HMI tags "Default tag table"
   "66_Event_Data_BC_EVENT_WORD_01" : Word = PLC "66_Event_Data".BC_EVENT_WORD_01 AT %DB66.DBW0, 1 s
   "66_Event_Data_BC_EVENT_WORD_02" : Word = PLC "66_Event_Data".BC_EVENT_WORD_02 AT %DB66.DBW2, 1 s
   "64_Message_Data_BC_MESSAGE_WORD_01" : Word = PLC "64_Message_Data".BC_MESSAGE_WORD_01 AT %DB64.DBW0, 1 s
   "64_Message_Data_BC_MESSAGE_WORD_02" : Word = PLC "64_Message_Data".BC_MESSAGE_WORD_02 AT %DB64.DBW2, 1 s
   "66_Event_Data_IGG_EVENT_WORD_01" : Word = PLC "66_Event_Data".IGG_EVENT_WORD_01 AT %DB66.DBW0, 1 s
   "66_Event_Data_IGG_EVENT_WORD_02" : Word = PLC "66_Event_Data".IGG_EVENT_WORD_02 AT %DB66.DBW2, 1 s
   "64_Message_Data_IGG_MESSAGE_WORD_01" : Word = PLC "64_Message_Data".IGG_MESSAGE_WORD_01 AT %DB64.DBW0, 1 s
   "64_Message_Data_IGG_MESSAGE_WORD_02" : Word = PLC "64_Message_Data".IGG_MESSAGE_WORD_02 AT %DB64.DBW2, 1 s
   "Current User" : WString[15] AT %DB1.DBX0.0
   "db_time_sync_time_system_READ" : LDT = PLC db_time_sync_time_system_READ AT %M2.0, 1 s
   "80_From_HMI_Cooling System Overrun" : Time = PLC "80_From_HMI"."Cooling System Overrun", 1 s
   "Start Sequenc_DB_Post Purge Time Sec" : Int, internal
   "db_time_sync_time_local_READ" : LDT = PLC db_time_sync_time_local_READ AT %M4.0, 1 s
   "82_To_HMI_Fuel Pump 1 Animation" : Int = PLC "82_To_HMI"."Fuel Pump 1 Animation", 1 s
   "82_To_HMI_Fuel Pump 2 Animation" : Int = PLC "82_To_HMI"."Fuel Pump 2 Animation", 1 s
   "16_AQ_Data_CV203_CNTRL(1)" : Real = PLC "16_AQ_Data".CV203_CNTRL, 1 s
   "HMI Data_O2 Setpoint" : Real, internal
   "82_To_HMI_IA Compressor Animation" : Int = PLC "82_To_HMI"."IA Compressor Animation", 1 s
   "Atomising Air  Valve Manual Regulator" : Int, internal
   "Fuel Valve Manual Regulator" : Int, internal
   "82_To_HMI_I&A Compressor Run Hours(1)" : Int = PLC "82_To_HMI"."I&A Compressor Run Hours", 1 s
   "82_To_HMI_I&A Compressor Service Time Hours" : Int = PLC "82_To_HMI"."I&A Compressor Service Time Hours", 1 s
   "82_To_HMI_CA Blower Run Days" : Int = PLC "82_To_HMI"."CA Blower Run Days", 1 s
   "82_To_HMI_CA Blower Service Time Hours" : Int = PLC "82_To_HMI"."CA Blower Service Time Hours", 1 s
   "82_To_HMI_CA Blower Run Hours" : Int = PLC "82_To_HMI"."CA Blower Run Hours", 1 s
   "82_To_HMI_CA Blower Run Minutes" : Int = PLC "82_To_HMI"."CA Blower Run Minutes", 1 s
   "82_To_HMI_I&A Compressor Run Minutes" : Int = PLC "82_To_HMI"."I&A Compressor Run Minutes", 1 s
   "82_To_HMI_I&A Compressor Run Seconds" : Int = PLC "82_To_HMI"."I&A Compressor Run Seconds", 1 s
   "P305_Functioning Hours_IDB_Hours Total" : Int = PLC "P305_Functioning Hours_IDB"."Hours Total", 1 s
   "82_To_HMI_P305 FW Pump Service Time Hours" : Int = PLC "82_To_HMI"."P305 FW Pump Service Time Hours", 1 s
   "P305_Functioning Hours_IDB_Service Time bit" : Bool = PLC "P305_Functioning Hours_IDB"."Service Time bit", 1 s
   "P305_Functioning Hours_IDB_Minutes" : Int = PLC "P305_Functioning Hours_IDB".Minutes, 1 s
   "P305_Functioning Hours_IDB_Seconds" : Int = PLC "20_TANKS_IP_DATA".RIO_04.SECOND_TANK.BWT_LEVEL_HIHI, 1 s
   "FW Pump Animation" : Int, internal
   "82_To_HMI_I&A Compressor Run Hours" : Int = PLC "82_To_HMI"."I&A Compressor Run Hours", 1 s
   "82_To_HMI_CRNT_MODE_IGG" : Int = PLC "82_To_HMI".CRNT_MODE_IGG, 1 s
   "70_Mode_Data_AUT_RST_PLS_IN" : Bool = PLC "70_Mode_Data".AUT_RST_PLS.IN, 1 s
   "RESET_STEP" : Bool = PLC RESET_STEP AT %M12.0, 1 s
   "100_IGG_AUTO_SEQ_DB_CRNT_STEP" : Int = PLC "100_IGG_AUTO_SEQ_DB".CRNT_STEP, 1 s
   "100_BC_AUTO_SEQ_DB_CRNT_STEP" : Int = PLC "100_BC_AUTO_SEQ_DB".CRNT_STEP, 1 s
   "103_Main_Burner_DB_RUN" : Bool = PLC "103_Main_Burner_DB".RUN, 1 s
   "60_Alarm_Data_ALRM_PRSNT" : Bool = PLC "60_Alarm_Data".ALRM_PRSNT AT %DB60.DBX32.0, 1 s
      on ChangeValue: "ALARM_Present"()
   "62_Warning_Data_WRNG_PRSNT" : Bool = PLC "62_Warning_Data".WRNG_PRSNT AT %DB62.DBX16.0, 1 s
   "103_Main_Burner_DB_RUNNING" : Bool = PLC "103_Main_Burner_DB".RUNNING, 1 s
   "101_Fuel_Pumps_DB_Duty Is B" : Bool = PLC "101_Fuel_Pumps_DB"."Duty Is B", 1 s
   "101_Fuel_Pumps_DB_Duty Is A" : Bool = PLC "101_Fuel_Pumps_DB"."Duty Is A", 1 s
   "84_Setpoints_PIT204_High" : Real = PLC "84_Setpoints".PIT204_High, 1 s
   "84_Setpoints_PIT204_High(1)" : Real = PLC "84_Setpoints".PIT204_High, 1 s
   "84_Setpoints_PIT204_HighHigh" : Real = PLC "84_Setpoints".PIT204_HighHigh, 1 s
   "84_Setpoints_PIT204_HighHigh(1)" : Real = PLC "84_Setpoints".PIT204_HighHigh, 1 s
   "84_Setpoints_PIT204_LowLow" : Real = PLC "84_Setpoints".PIT204_LowLow, 1 s
   "84_Setpoints_PIT204_LowLow(1)" : Real = PLC "84_Setpoints".PIT204_LowLow, 1 s
   "84_Setpoints_PIT204_Low" : Real = PLC "84_Setpoints".PIT204_Low, 1 s
   "84_Setpoints_PIT204_Low(1)" : Real = PLC "84_Setpoints".PIT204_Low, 1 s
   "80_From_HMI_RST_LOCKOUT" : Bool = PLC "80_From_HMI".RST_LOCKOUT, 1 s
   "80_From_HMI_Beacon frequency" : Time = PLC "80_From_HMI"."Beacon frequency", 1 s
   "80_From_HMI_Buzzer reset time" : Time = PLC "80_From_HMI"."Buzzer reset time", 1 s
   "80_From_HMI_Reset_Alarms" : Bool = PLC "80_From_HMI".Reset_Alarms, 1 s
   "Alarm beacon handling_DB_Buzzer_Timer_0_Instance_Q" : Bool = PLC "Alarm beacon handling_DB".Buzzer_Timer_0_Instance.Q, 1 s
   "Buzzer" : Bool = PLC Buzzer AT %Q1.7, 1 s
   "80_From_HMI_FLM_FAIL_DLY" : Time = PLC "80_From_HMI".FLM_FAIL_DLY, 1 s
   "103_Main_Burner_DB_DN_OK" : Bool = PLC "103_Main_Burner_DB".DN_OK, 1 s
   "103_Main_Burner_DB_Days burn_CV" : Int = PLC "103_Main_Burner_DB"."Days burn".CV, 1 s
   "103_Main_Burner_DB_Hours burn_CV" : Int = PLC "103_Main_Burner_DB"."Hours burn".CV, 1 s
   "103_Main_Burner_DB_Minutes burn_CV" : Int = PLC "103_Main_Burner_DB"."Minutes burn".CV, 1 s
   "103_Main_Burner_DB_Seconds burn_CV" : Int = PLC "103_Main_Burner_DB"."Seconds burn".CV, 1 s
   "103_Main_Burner_DB_STATE" : Int = PLC "103_Main_Burner_DB".STATE, 1 s
   "19_AUTO_CMNDS_Data_CV203_RAMP_CNTRL" : Bool = PLC "19_AUTO_CMNDS_Data".CV203_RAMP_CNTRL, 1 s
   "102_Pilot_Burner_DB_RUNNING" : Bool = PLC "102_Pilot_Burner_DB".RUNNING, 1 s
   "68_Sys_Status_Data_FUEL_PRES_IN_RNG" : Bool = PLC "68_Sys_Status_Data".FUEL_PRES_IN_RNG, 1 s
   "68_Sys_Status_Data_IA_PRES_IN_RNG" : Bool = PLC "68_Sys_Status_Data".IA_PRES_IN_RNG, 1 s
   "84_Setpoints_Gain" : Real = PLC "84_Setpoints".Gain, 1 s
   "84_Setpoints_Integration Time" : Time = PLC "84_Setpoints"."Integration Time", 1 s
   "84_Setpoints_Derive Time" : Time = PLC "84_Setpoints"."Derive Time", 1 s
   "O2 Ramp Control_QLMN_HLM" : Bool = PLC "O2 Ramp Control".QLMN_HLM, 1 s
   "O2 Ramp Control_QLMN_LLM" : Bool = PLC "O2 Ramp Control".QLMN_LLM, 1 s
   "84_Setpoints_P_ON" : Bool = PLC "84_Setpoints".P_ON, 1 s
   "84_Setpoints_I_ON" : Bool = PLC "84_Setpoints".I_ON, 1 s
   "84_Setpoints_D_ON" : Bool = PLC "84_Setpoints".D_ON, 1 s
   "Evolving Setpoint_DB_LevelBetter" : Bool = PLC "Evolving Setpoint_DB".LevelBetter, 1 s
   "84_Setpoints_Max Opening" : Real = PLC "84_Setpoints"."Max Opening", 1 s
   "84_Setpoints_Min Opening" : Real = PLC "86_Times".STEP_MAX_TIME_STP_290, 1 s
   "80_From_HMI_Post Purge Time" : Time = PLC "80_From_HMI"."Post Purge Time", 1 s
   "103_Main_Burner_DB_Status" : Int = PLC "103_Main_Burner_DB".Status, 1 s
   "80_From_HMI_Reset CV203 PID" : Bool = PLC "80_From_HMI"."Reset CV203 PID", 1 s
   "80_From_HMI_BurnerProgramedStop" : Bool = PLC "80_From_HMI".BurnerProgramedStop, 1 s
   "82_To_HMI_CA Blower Reset Hours" : Bool = PLC "82_To_HMI"."CA Blower Reset Hours", 1 s
   "82_To_HMI_CA Blower Service Due" : Bool = PLC "82_To_HMI"."CA Blower Service Due", 1 s
   "Operation hours E139_IDB_Hours Functioning" : Int = PLC "Operation hours E139_IDB"."Hours Functioning", 1 s
   "82_To_HMI_CA Blower Total Run Hours" : Int = PLC "82_To_HMI"."CA Blower Total Run Hours", 1 s
   "82_To_HMI_I&A Compressor Total Run Hours" : Int = PLC "82_To_HMI"."I&A Compressor Total Run Hours", 1 s
   "82_To_HMI_I&A Compressor Reset Hours" : Bool = PLC "82_To_HMI"."I&A Compressor Reset Hours", 1 s
   "82_To_HMI_I&A Compressor Service Due" : Bool = PLC "82_To_HMI"."I&A Compressor Service Due", 1 s
   "82_To_HMI_E500A Fuel Pump Run Hours" : Int = PLC "82_To_HMI"."E500A Fuel Pump Run Hours", 1 s
   "64_Functioning Hours_E500A_IDB_Hours Functioning" : Int = PLC "64_Functioning Hours_E500A_IDB"."Hours Functioning", 1 s
   "82_To_HMI_E500A Fuel Pump Run Minutes" : Int = PLC "82_To_HMI"."E500A Fuel Pump Run Minutes", 1 s
   "82_To_HMI_E500A Fuel Pump Run Seconds" : Int = PLC "82_To_HMI"."E500A Fuel Pump Run Seconds", 1 s
   "82_To_HMI_E500A Fuel Pump Total Run Hours" : Int = PLC "82_To_HMI"."E500A Fuel Pump Total Run Hours", 1 s
   "82_To_HMI_E500A Fuel Pump Service Time Hours" : Int = PLC "82_To_HMI"."E500A Fuel Pump Service Time Hours", 1 s
   "82_To_HMI_E500A Fuel Pump Reset Hours" : Bool = PLC "82_To_HMI"."E500A Fuel Pump Reset Hours", 1 s
   "64_Functioning Hours_E500B_IDB_Hours Functioning" : Int = PLC "64_Functioning Hours_E500B_IDB"."Hours Functioning", 1 s
   "82_To_HMI_E500B Fuel Pump Run Minutes" : Int = PLC "82_To_HMI"."E500B Fuel Pump Run Minutes", 1 s
   "82_To_HMI_E500B Fuel Pump Run Seconds" : Int = PLC "82_To_HMI"."E500B Fuel Pump Run Seconds", 1 s
   "82_To_HMI_E500B Fuel Pump Total Run Hours" : Int = PLC "82_To_HMI"."E500B Fuel Pump Total Run Hours", 1 s
   "82_To_HMI_E500B Fuel Pump Service Time Hours" : Int = PLC "82_To_HMI"."E500B Fuel Pump Service Time Hours", 1 s
   "82_To_HMI_E500B Fuel Pump Reset Hours" : Bool = PLC "82_To_HMI"."E500B Fuel Pump Reset Hours", 1 s
   "82_To_HMI_E500B Fuel Pump Service Due" : Bool = PLC "82_To_HMI"."E500B Fuel Pump Service Due", 1 s
   "82_To_HMI_E500A Fuel Pump Service Due" : Bool = PLC "82_To_HMI"."E500A Fuel Pump Service Due", 1 s
   "64_Functioning Hours_P301_IDB_Hours Functioning" : Int = PLC "64_Functioning Hours_P301_IDB"."Hours Functioning", 1 s
   "82_To_HMI_P301 CSW Pump Run Minutes" : Int = PLC "82_To_HMI"."P301 CSW Pump Run Minutes", 1 s
   "82_To_HMI_P301 CSW Pump Run Seconds" : Int = PLC "82_To_HMI"."P301 CSW Pump Run Seconds", 1 s
   "82_To_HMI_P301 CSW Pump Reset Hours" : Bool = PLC "82_To_HMI"."P301 CSW Pump Reset Hours", 1 s
   "82_To_HMI_P301 CSW Pump Service Due" : Bool = PLC "82_To_HMI"."P301 CSW Pump Service Due", 1 s
   "80_From_HMI_P301_PRSNT" : Bool = PLC "80_From_HMI".P301_PRSNT, 1 s
   "Alarms_Acknowledge_IGG_ALARM_ACKNLG_3" : Word = PLC Alarms_Acknowledge.IGG_ALARM_ACKNLG_3 AT %DB67.DBW4, 1 s
   "Alarms_Acknowledge_IGG_ALARM_ACKNLG_4" : Word = PLC Alarms_Acknowledge.IGG_ALARM_ACKNLG_4 AT %DB67.DBW6, 1 s
   "Alarms_Acknowledge_IGG_ALARM_ACKNLG_2" : Word = PLC Alarms_Acknowledge.IGG_ALARM_ACKNLG_2 AT %DB67.DBW2, 1 s
   "Alarms_Acknowledge_IGG_ALARM_ACKNLG_1" : Word = PLC Alarms_Acknowledge.IGG_ALARM_ACKNLG_1 AT %DB67.DBW0, 1 s
   "BC_ALARM_ACKNLG_1" : Word = PLC BC_ALARM_ACKNLG_1 AT %MW24, 1 s
   "BC_ALARM_ACKNLG_2" : Word = PLC BC_ALARM_ACKNLG_2 AT %MW26, 1 s
   "BC_ALARM_ACKNLG_3" : Word = PLC BC_ALARM_ACKNLG_3 AT %MW28, 1 s
   "BC_ALARM_ACKNLG_4" : Word = PLC BC_ALARM_ACKNLG_4 AT %MW30, 1 s
   "80_From_HMI_P305_PRSNT" : Bool = PLC "80_From_HMI".P305_PRSNT, 1 s
   "68_Sys_Status_Data_INTRLKS_OK" : Bool = PLC "68_Sys_Status_Data".INTRLKS_OK, 1 s
   "82_To_HMI_E-STOP LATCHED" : Bool = PLC "82_To_HMI"."E-STOP LATCHED", 1 s
   "82_To_HMI_P301 CSW Pump Run Days" : Int = PLC "82_To_HMI"."P301 CSW Pump Run Days", 1 s
   "82_To_HMI_CA Blower Run Seconds" : Int = PLC "82_To_HMI"."CA Blower Run Seconds", 1 s
   "82_To_HMI_P305 FW Pump Reset Hours" : Bool = PLC "82_To_HMI"."P305 FW Pump Reset Hours", 1 s
   "P305_Functioning Hours_IDB_Hours Functioning Out" : Int = PLC "P305_Functioning Hours_IDB"."Hours Functioning Out", 1 s
   "82_To_HMI_P305 FW Pump Run Hours" : Int = PLC "82_To_HMI"."P305 FW Pump Run Hours", 1 s
   "82_To_HMI_P305 FW Pump Run Days" : Int = PLC "82_To_HMI"."P305 FW Pump Run Days", 1 s
   "82_To_HMI_P301 CSW Pump Service Time Hours" : Int = PLC "82_To_HMI"."P301 CSW Pump Service Time Hours", 1 s
   "82_To_HMI_P301 CSW Pump Run Hours" : Int = PLC "82_To_HMI"."P301 CSW Pump Run Hours", 1 s
   "82_To_HMI_P301 CSW Pump Total Run Hours" : Int = PLC "82_To_HMI"."P301 CSW Pump Total Run Hours", 1 s
   "80_From_HMI_PIT 359 delay" : Time = PLC "80_From_HMI"."PIT 359 delay", 1 s
   "80_From_HMI_PIT 316 delay" : Time = PLC "80_From_HMI"."PIT 316 delay", 1 s
   "86_Times_PIT353 Delay" : Time = PLC "86_Times"."PIT353 Delay", 1 s
   "86_Times_PIT416 Delay" : Time = PLC "86_Times"."PIT416 Delay", 1 s
   "19_AUTO_CMNDS_Data_PIT416_CMND_Target" : Real = PLC "19_AUTO_CMNDS_Data".PIT416_CMND_Target, 1 s
   "2102_TIME_CALCS_DB_Voyage_TIME_days" : Int = PLC "2102_TIME_CALCS_DB".Voyage_TIME_days, 1 s
   "2102_TIME_CALCS_DB_Voyage_TIME_invalid" : Bool = PLC "2102_TIME_CALCS_DB".Voyage_TIME_invalid AT %DB1.DBW0, 1 s
      on ChangeValue: "VoyageTimeInsufficient"()
   "2102_TIME_CALCS_DB_TOT_SEQ_DAYS" : Real = PLC "2102_TIME_CALCS_DB".TOT_SEQ_DAYS, 1 s
   "2102_TIME_CALCS_DB_POST_DWELL_TMR_DN(1)" : Bool = PLC "2102_TIME_CALCS_DB".POST_DWELL_TMR_DN AT %DB1.DBD0, 1 s
   "2102_TIME_CALCS_DB_PRE-DWEL HOURS REMNG" : Int = PLC "2102_TIME_CALCS_DB"."PRE-DWEL HOURS REMNG" AT %DB1.DBW0, 1 s
   "504_Tank Grouping_DB2020_TANK ACTIV 2" : Bool = PLC "504_Tank Grouping_DB2020"."TANK ACTIV 2" AT %DB1.DBW0, 1 s
   "504_Tank Grouping_DB2020_TANK ACTIV 4" : Bool = PLC "504_Tank Grouping_DB2020"."TANK ACTIV 4" AT %DB1.DBW0, 1 s
   "504_Tank Grouping_DB2020_TANK ACTIV 6" : Bool = PLC "504_Tank Grouping_DB2020"."TANK ACTIV 6" AT %DB1.DBW0, 1 s
   "504_Tank Grouping_DB2020_TANK ACTIV 8" : Bool = PLC "504_Tank Grouping_DB2020"."TANK ACTIV 8" AT %DB1.DBW0, 1 s
   "504_Tank Grouping_DB2020_TANK ACTIV 10" : Bool = PLC "504_Tank Grouping_DB2020"."TANK ACTIV 10" AT %DB1.DBW0, 1 s
   "504_Tank Grouping_DB2020_TANK ACTIV 12" : Bool = PLC "504_Tank Grouping_DB2020"."TANK ACTIV 12" AT %DB1.DBW0, 1 s
   "504_Tank Grouping_DB2020_TANK ACTIV 14" : Bool = PLC "504_Tank Grouping_DB2020"."TANK ACTIV 14" AT %DB1.DBW0, 1 s
   "504_Tank Grouping_DB2020_TANK ACTIV 16" : Bool = PLC "504_Tank Grouping_DB2020"."TANK ACTIV 16" AT %DB1.DBW0, 1 s
   "504_Tank Grouping_DB2020_TANK ACTIV 18" : Bool = PLC "504_Tank Grouping_DB2020"."TANK ACTIV 18" AT %DB1.DBW0, 1 s
   "504_Tank Grouping_DB2020_TANK ACTIV 20" : Bool = PLC "504_Tank Grouping_DB2020"."TANK ACTIV 20" AT %DB1.DBW0, 1 s
   "504_Tank Grouping_DB2020_TANK ACTIV 3" : Bool = PLC "504_Tank Grouping_DB2020"."TANK ACTIV 3" AT %DB1.DBW0, 1 s
   "504_Tank Grouping_DB2020_TANK ACTIV 5" : Bool = PLC "504_Tank Grouping_DB2020"."TANK ACTIV 5" AT %DB1.DBW0, 1 s
   "504_Tank Grouping_DB2020_TANK ACTIV 7" : Bool = PLC "504_Tank Grouping_DB2020"."TANK ACTIV 7" AT %DB1.DBW0, 1 s
   "504_Tank Grouping_DB2020_TANK ACTIV 9" : Bool = PLC "504_Tank Grouping_DB2020"."TANK ACTIV 9" AT %DB1.DBW0, 1 s
   "504_Tank Grouping_DB2020_TANK ACTIV 11" : Bool = PLC "504_Tank Grouping_DB2020"."TANK ACTIV 11" AT %DB1.DBW0, 1 s
   "504_Tank Grouping_DB2020_TANK ACTIV 13" : Bool = PLC "504_Tank Grouping_DB2020"."TANK ACTIV 13" AT %DB1.DBW0, 1 s
   "504_Tank Grouping_DB2020_TANK ACTIV 1" : Bool = PLC "504_Tank Grouping_DB2020"."TANK ACTIV 1" AT %DB1.DBW0, 1 s
   "504_Tank Grouping_DB2020_TANK ACTIV 17" : Bool = PLC "504_Tank Grouping_DB2020"."TANK ACTIV 17" AT %DB1.DBW0, 1 s
   "504_Tank Grouping_DB2020_TANK ACTIV 19" : Bool = PLC "504_Tank Grouping_DB2020"."TANK ACTIV 19" AT %DB1.DBW0, 1 s
   "504_Tank Grouping_DB2020_TANK ACTIV 21" : Bool = PLC "504_Tank Grouping_DB2020"."TANK ACTIV 21" AT %DB1.DBW0, 1 s
   "2110_BTCS_CNTRL_DB_PORT_TANK_STS(1)" : Bool = PLC "2110_BTCS_CNTRL_DB".PORT_TANK_STS AT %DB1.DBX0.0, 1 s
   "Tank Activated Port 2" : Int, internal
   "Tank Activated Port 3" : Int, internal
   "Tank Activated Port 4" : Int, internal
   "Tank Activated Port 5" : Int, internal
   "Tank Activated Port 6" : Int, internal
   "Tank Activated Port 7" : Int, internal
   "Tank Activated Port 8" : Int, internal
   "Tank Activated Port 9" : Int, internal
   "Tank Activated Port 10" : Int, internal
   "2110_BTCS_CNTRL_DB_STBD_TANK_STS(1)" : Bool = PLC "20_TANKS_IP_DATA".RIO_01.FIRST_TANK.GTT_ISOL_VALVE_OPEN, 1 s
   "Tank Activated Star 2" : Int, internal
   "Tank Activated Star 3" : Int, internal
   "Tank Activated Star 4" : Int, internal
   "Tank Activated Star 5" : Int, internal
   "Tank Activated Star 6" : Int, internal
   "Tank Activated Star 7" : Int, internal
   "Tank Activated Star 8" : Int, internal
   "Tank Activated Star 9" : Int, internal
   "Tank Activated Star 10" : Int, internal
   "2102_TIME_CALCS_DB_PRE-DWEL_Warning 1" : Bool = PLC "2102_TIME_CALCS_DB"."PRE-DWEL_Warning 1", 500 ms
      on ChangeValue: "TimeRemainingToTreatment"()
   "2102_TIME_CALCS_DB_PRE-DWEL_Warning Min 1" : Int = PLC "2102_TIME_CALCS_DB"."PRE-DWEL_Warning Min 1", 1 s
   "2102_TIME_CALCS_DB_PRE-DWEL_Warning Min 2" : Int = PLC "2102_TIME_CALCS_DB"."PRE-DWEL_Warning Min 2", 1 s
   "2102_TIME_CALCS_DB_PRE-DWEL_Warning Min 3" : Int = PLC "2102_TIME_CALCS_DB"."PRE-DWEL_Warning Min 3", 1 s
   "2102_TIME_CALCS_DB_PRE-DWEL_Warning Reset 1" : Bool = PLC "2102_TIME_CALCS_DB"."PRE-DWEL_Warning Reset 1", 1 s
   "2102_TIME_CALCS_DB_PRE-DWEL_Warning 2" : Bool = PLC "2102_TIME_CALCS_DB"."PRE-DWEL_Warning 2", 500 ms
      on ChangeValue: "TreatmentRequired"()
   "2102_TIME_CALCS_DB_PRE-DWEL_Warning 3" : Bool = PLC "2102_TIME_CALCS_DB"."PRE-DWEL_Warning 3", 1 s
   "2102_TIME_CALCS_DB_PRE-DWEL_Warning Reset 2" : Bool = PLC "2102_TIME_CALCS_DB"."PRE-DWEL_Warning Reset 2", 1 s
   "2102_TIME_CALCS_DB_PRE-DWEL_Warning Reset 3" : Bool = PLC "2102_TIME_CALCS_DB"."PRE-DWEL_Warning Reset 3", 1 s
   "2102_TIME_CALCS_DB_60X boost" : Bool = PLC "2102_TIME_CALCS_DB"."60X boost", 1 s
   "86_Times_P301_START_DLY" : Time = PLC "86_Times".P301_START_DLY, 1 s
   "86_Times_FS332 Delay" : Time = PLC "86_Times"."FS332 Delay", 1 s
   "86_Times_LIT304 Delay" : Time = PLC "86_Times"."LIT304 Delay", 1 s
   "86_Times_PIT402_Ramp_Seconds" : Int = PLC "86_Times".PIT402_Ramp_Seconds, 1 s
   "86_Times_PIT402 Alarm Delay" : Time = PLC "86_Times"."PIT402 Alarm Delay", 1 s
   "84_Setpoints_PIT113_Burner_Target" : Real = PLC "84_Setpoints".PIT113_Burner_Target, 1 s
   "2102_TIME_CALCS_DB_PRE-DWEL MINS REMNG" : Int = PLC "2102_TIME_CALCS_DB"."PRE-DWEL MINS REMNG", 1 s
   "84_Setpoints_LIT304_InitialFill_Target_Low" : Real = PLC "84_Setpoints".LIT304_InitialFill_Target_Low, 1 s
   "84_Setpoints_LIT304_Refill_Target_Low" : Real = PLC "84_Setpoints".LIT304_Refill_Target_Low, 1 s
   "1111_PID_CV111_Setpoint" : Real = PLC "1111_PID_CV111".Setpoint, 1 s
   "2086_Times_TT426_PORT_Alarm Delay" : Time = PLC "2086_Times"."TT426_PORT_Alarm Delay", 1 s
   "2086_Times_TT426_STAR_Alarm Delay" : Time = PLC "2086_Times"."TT426_STAR_Alarm Delay", 1 s
   "2086_Times_FIT418PORT Alarm Delay" : Time = PLC "2086_Times"."FIT418PORT Alarm Delay", 1 s
   "2086_Times_FIT420PORT Alarm Delay" : Time = PLC "2086_Times"."FIT420PORT Alarm Delay", 1 s
   "2086_Times_FIT417STAR Alarm Delay" : Time = PLC "2086_Times"."FIT417STAR Alarm Delay", 1 s
   "2086_Times_FIT419STAR Alarm Delay" : Time = PLC "2086_Times"."FIT419STAR Alarm Delay", 1 s
   "2086_Times_PT415 Alarm Delay" : Time = PLC "2086_Times"."PT415 Alarm Delay", 1 s
   "2086_Times_PIT424 Alarm Delay" : Time = PLC "2086_Times"."PIT424 Alarm Delay", 1 s
   "2086_Times_LS425 Port Alarm Delay" : Time = PLC "2086_Times"."LS425 Port Alarm Delay", 1 s
   "2086_Times_LS425 Star Alarm Delay" : Time = PLC "2086_Times"."LS425 Star Alarm Delay", 1 s
   "2086_Times_PS436 Alarm Delay" : Time = PLC "2086_Times"."PS436 Alarm Delay", 1 s
   "2102_TIME_CALCS_DB_Voyage_TIME_remaining_m" : Int = PLC "2102_TIME_CALCS_DB".Voyage_TIME_remaining_m, 1 s
   "2102_TIME_CALCS_DB_Voyage_TIME_remaining_h" : Int = PLC "2102_TIME_CALCS_DB".Voyage_TIME_remaining_h, 1 s
   "2102_TIME_CALCS_DB_Time_To_Treatment" : Int = PLC "2102_TIME_CALCS_DB".Time_To_Treatment, 1 s
   "PGC_COMMISSION_MODE_DB_Setpoint" : Real = PLC PGC_COMMISSION_MODE_DB.Setpoint, 1 s
   "PGC_COMMISSION_MODE_DB_Button Control" : Int = PLC PGC_COMMISSION_MODE_DB."Button Control", 1 s
   "PGC_COMMISSION_MODE_DB_Active" : Bool = PLC PGC_COMMISSION_MODE_DB.Active, 1 s
   "PGC_COMMISSION_MODE_DB_Drive Popup" : Bool = PLC PGC_COMMISSION_MODE_DB."Drive Popup", 500 ms
      on ChangeValue: "PGCCommissioning"()
   "21_FLOW_PRESSURE_SETPOINT_FIT_419_PRESSURE_SETPOINT" : Real = PLC "21_FLOW_PRESSURE_SETPOINT".FIT_419_PRESSURE_SETPOINT, 1 s
   "21_FLOW_PRESSURE_SETPOINT_FIT_420_PRESSURE_SETPOINT" : Real = PLC "21_FLOW_PRESSURE_SETPOINT".FIT_420_PRESSURE_SETPOINT, 1 s
   "user_group" : Int, internal
   "2102_TIME_CALCS_DB_Voyage_TIME_hours" : Int = PLC "2102_TIME_CALCS_DB".Voyage_TIME_hours, 1 s
   "2115_VOYAGE_TIME_DAYS_VOYAGE_DAYS" : Real = PLC "2115_VOYAGE_TIME_DAYS".VOYAGE_DAYS, 1 s
   "2102_TIME_CALCS_DB_PHASE_DIFFERECE_MNS_REMNG_De-Ox" : Int = PLC "2102_TIME_CALCS_DB".PHASE_DIFFERECE_MNS_REMNG_De-Ox, 1 s
   "504_Tank Grouping_DB2020_SetGroup" : Bool = PLC "2060_Alarm_Data".BTCS_ALARM_WORD_05, 1 s
   "504_Tank Grouping_DB2020_GROUP of TANK 1" : Int = PLC "504_Tank Grouping_DB2020"."GROUP of TANK 1", 1 s
   "504_Tank Grouping_DB2020_GROUP of TANK 2" : Int = PLC "504_Tank Grouping_DB2020"."GROUP of TANK 2", 1 s
   "504_Tank Grouping_DB2020_GROUP of TANK 3" : Int = PLC "504_Tank Grouping_DB2020"."GROUP of TANK 3", 1 s
   "504_Tank Grouping_DB2020_GROUP of TANK 4" : Int = PLC "504_Tank Grouping_DB2020"."GROUP of TANK 4", 1 s
   "504_Tank Grouping_DB2020_GROUP of TANK 5" : Int = PLC "504_Tank Grouping_DB2020"."GROUP of TANK 5", 1 s
   "504_Tank Grouping_DB2020_GROUP of TANK 6" : Int = PLC "504_Tank Grouping_DB2020"."GROUP of TANK 6", 1 s
   "504_Tank Grouping_DB2020_GROUP of TANK 7" : Int = PLC "504_Tank Grouping_DB2020"."GROUP of TANK 7", 1 s
   "504_Tank Grouping_DB2020_GROUP of TANK 8" : Int = PLC "504_Tank Grouping_DB2020"."GROUP of TANK 8", 1 s
   "504_Tank Grouping_DB2020_GROUP of TANK 9" : Int = PLC "504_Tank Grouping_DB2020"."GROUP of TANK 9", 1 s
   "504_Tank Grouping_DB2020_GROUP of TANK 10" : Int = PLC "504_Tank Grouping_DB2020"."GROUP of TANK 10", 1 s
   "504_Tank Grouping_DB2020_GROUP of TANK 11" : Int = PLC "504_Tank Grouping_DB2020"."GROUP of TANK 11", 1 s
   "504_Tank Grouping_DB2020_GROUP of TANK 12" : Int = PLC "504_Tank Grouping_DB2020"."GROUP of TANK 12", 1 s
   "504_Tank Grouping_DB2020_GROUP of TANK 13" : Int = PLC "504_Tank Grouping_DB2020"."GROUP of TANK 13", 1 s
   "504_Tank Grouping_DB2020_GROUP of TANK 14" : Int = PLC "504_Tank Grouping_DB2020"."GROUP of TANK 14", 1 s
   "504_Tank Grouping_DB2020_GROUP ACTIV 1" : Bool = PLC "504_Tank Grouping_DB2020"."GROUP ACTIV 1", 1 s
   "504_Tank Grouping_DB2020_GROUP ACTIV 2" : Bool = PLC "504_Tank Grouping_DB2020"."GROUP ACTIV 2", 1 s
   "504_Tank Grouping_DB2020_GROUP ACTIV 3" : Bool = PLC "504_Tank Grouping_DB2020"."GROUP ACTIV 3", 1 s
   "504_Tank Grouping_DB2020_GROUP ACTIV 4" : Bool = PLC "504_Tank Grouping_DB2020"."GROUP ACTIV 4", 1 s
   "504_Tank Grouping_DB2020_GROUP ACTIV 5" : Bool = PLC "504_Tank Grouping_DB2020"."GROUP ACTIV 5", 1 s
   "504_Tank Grouping_DB2020_GROUP ACTIV 6" : Bool = PLC "504_Tank Grouping_DB2020"."GROUP ACTIV 6", 1 s
   "504_Tank Grouping_DB2020_GROUP ACTIV 7" : Bool = PLC "504_Tank Grouping_DB2020"."GROUP ACTIV 7", 1 s
   "504_Tank Grouping_DB2020_GROUP SET" : Int = PLC "504_Tank Grouping_DB2020"."GROUP SET", 1 s
   "504_Tank Grouping_DB2020_GROUP ACTIVE INT 1" : Bool = PLC "504_Tank Grouping_DB2020"."GROUP ACTIVE INT 1", 1 s
   "504_Tank Grouping_DB2020_GROUP ACTIVE INT 2" : Bool = PLC "504_Tank Grouping_DB2020"."GROUP ACTIVE INT 2", 1 s
   "504_Tank Grouping_DB2020_GROUP ACTIVE INT 3" : Bool = PLC "504_Tank Grouping_DB2020"."GROUP ACTIVE INT 3", 1 s
   "504_Tank Grouping_DB2020_GROUP ACTIVE INT 4" : Bool = PLC "504_Tank Grouping_DB2020"."GROUP ACTIVE INT 4", 1 s
   "504_Tank Grouping_DB2020_GROUP ACTIVE INT 5" : Bool = PLC "504_Tank Grouping_DB2020"."GROUP ACTIVE INT 5", 1 s
   "504_Tank Grouping_DB2020_GROUP ACTIVE INT 6" : Bool = PLC "504_Tank Grouping_DB2020"."GROUP ACTIVE INT 6", 1 s
   "504_Tank Grouping_DB2020_GROUP ACTIVE INT 7" : Bool = PLC "504_Tank Grouping_DB2020"."GROUP ACTIVE INT 7", 1 s
   "80_From_HMI_TIMER RST Supres" : Bool = PLC "80_From_HMI"."TIMER RST Supres", 1 s
   "HMI Indication Logic_DB_FA Mode Selected" : Bool = PLC "HMI Indication Logic_DB"."FA Mode Selected", 1 s
   "HMI Indication Logic_DB_Tank Selected" : Bool = PLC "HMI Indication Logic_DB"."Tank Selected", 1 s
   "51_SLAVE_STATUS_RUNNING" : Bool = PLC "51_SLAVE_STATUS".RUNNING AT %DB51.DBX4.2, 1 s
      on ChangeValue: function_fd9437ed(0, "IGG_BC_FD001_Flame Detector"); function_fd9437ed(0, "GCU_FW_TIT408_Fresh water cooling"); function_fd9437ed(0, "IGG_Fuel_TIT202_Fuel Oil"); function_fd9437ed(0, "IGG_IG_TIT401_IG vent"); function_fd9437ed(0, "IGG_SW_TIT319_Cooling water (main line)"); function_fd9437ed(0, "IGG_SW_TIT360_Cooling water to drain line"); function_fd9437ed(0, "IGG_SW_TIT315_CW Temp to IGG Jacket"); function_fd9437ed(0, "IGG_CAB_PIT102_Comb Air"); function_fd9437ed(0, "IGG_Fuel_PIT204_Fuel Oil"); function_fd9437ed(0, "IGG_IA_PIT113_Atom Air to MBurner"); function_fd9437ed(0, "IGG_Fuel_PIT205_Fuel to MBurner"); function_fd9437ed(0, "IGG_IG_PIT402_IG vent"); function_fd9437ed(0, "IGG_SW_PIT359_Cooling water (main line)"); function_fd9437ed(0, "IGG_IA_PIT112_Inst Air"); function_fd9437ed(0, "IGG_SW_PIT316_Cooling water to IGG Jacket"); function_fd9437ed(0, "IGG_IG_TX-431_Atm Oxygen 1")
   "HMI Indication Logic_DB_Sequence Finished" : Bool = PLC "HMI Indication Logic_DB"."Sequence Finished", 1 s
   "20_TANKS_IP_DATA_RIO_01_FIRST_TANK_BWT_LEVEL_HIHI" : Bool = PLC "20_TANKS_IP_DATA".RIO_01.FIRST_TANK.BWT_LEVEL_HIHI, 1 s
   "20_TANKS_IP_DATA_RIO_01_FIRST_TANK_MBG_FLOW" : Real = PLC "20_TANKS_IP_DATA".RIO_01.FIRST_TANK.MBG_FLOW, 1 s
   "20_TANKS_IP_DATA_RIO_01_FIRST_TANK_USD_FLOW" : Real = PLC "20_TANKS_IP_DATA".RIO_01.FIRST_TANK.USD_FLOW, 1 s
   "20_TANKS_IP_DATA_RIO_01_FIRST_TANK_GTT_ISOL_VALVE_OPEN" : Bool = PLC "20_TANKS_IP_DATA".RIO_01.FIRST_TANK.GTT_ISOL_VALVE_OPEN, 1 s
   "504_Tank Grouping_DB2020_RUN TANK 1" : Bool = PLC "504_Tank Grouping_DB2020"."RUN TANK 1", 1 s
   "504_Tank Grouping_DB2020_RUN TANK 2" : Bool = PLC "504_Tank Grouping_DB2020"."RUN TANK 2", 1 s
   "20_TANKS_IP_DATA_RIO_01_SECOND_TANK_BWT_LEVEL_HIHI" : Bool = PLC "20_TANKS_IP_DATA".RIO_01.SECOND_TANK.BWT_LEVEL_HIHI, 1 s
   "20_TANKS_IP_DATA_RIO_01_SECOND_TANK_USD_FLOW" : Real = PLC "20_TANKS_IP_DATA".RIO_01.SECOND_TANK.USD_FLOW, 1 s
   "20_TANKS_IP_DATA_RIO_01_SECOND_TANK_MBG_FLOW" : Real = PLC PGC_COMMISSION_MODE_DB."Button Control", 1 s
   "20_TANKS_IP_DATA_RIO_01_SECOND_TANK_GTT_ISOL_VALVE_OPEN" : Bool = PLC "20_TANKS_IP_DATA".RIO_01.SECOND_TANK.GTT_ISOL_VALVE_OPEN, 1 s
   "20_TANKS_IP_DATA_RIO_01_SECOND_TANK_GTT_ISOL_VALVE_CLSD" : Bool = PLC "20_TANKS_IP_DATA".RIO_01.SECOND_TANK.GTT_ISOL_VALVE_CLSD, 1 s
   "20_TANKS_IP_DATA_RIO_01_FIRST_TANK_GTT_ISOL_VALVE_CLSD" : Bool = PLC "20_TANKS_IP_DATA".RIO_01.FIRST_TANK.GTT_ISOL_VALVE_CLSD, 1 s
   "20_TANKS_IP_DATA_RIO_01_THIRD_TANK_BWT_LEVEL_HIHI" : Bool = PLC "20_TANKS_IP_DATA".RIO_01.THIRD_TANK.BWT_LEVEL_HIHI, 1 s
   "504_Tank Grouping_DB2020_RUN TANK 3" : Bool = PLC "504_Tank Grouping_DB2020"."RUN TANK 3", 1 s
   "20_TANKS_IP_DATA_RIO_01_THIRD_TANK_USD_FLOW" : Real = PLC "20_TANKS_IP_DATA".RIO_01.THIRD_TANK.USD_FLOW, 1 s
   "20_TANKS_IP_DATA_RIO_01_THIRD_TANK_MBG_FLOW" : Real = PLC "20_TANKS_IP_DATA".RIO_01.THIRD_TANK.MBG_FLOW, 1 s
   "20_TANKS_IP_DATA_RIO_01_THIRD_TANK_GTT_ISOL_VALVE_OPEN" : Bool = PLC "20_TANKS_IP_DATA".RIO_01.THIRD_TANK.GTT_ISOL_VALVE_OPEN, 1 s
   "20_TANKS_IP_DATA_RIO_01_THIRD_TANK_GTT_ISOL_VALVE_CLSD" : Bool = PLC "20_TANKS_IP_DATA".RIO_01.THIRD_TANK.GTT_ISOL_VALVE_CLSD, 1 s
   "504_Tank Grouping_DB2020_RUN TANK 4" : Bool = PLC "504_Tank Grouping_DB2020"."RUN TANK 4", 1 s
   "504_Tank Grouping_DB2020_RUN TANK 5" : Bool = PLC "504_Tank Grouping_DB2020"."RUN TANK 5", 1 s
   "20_TANKS_IP_DATA_RIO_03_FIRST_TANK_MBG_FLOW" : Real = PLC "20_TANKS_IP_DATA".RIO_03.FIRST_TANK.MBG_FLOW, 1 s
   "20_TANKS_IP_DATA_RIO_03_FIRST_TANK_USD_FLOW" : Real = PLC "20_TANKS_IP_DATA".RIO_03.FIRST_TANK.USD_FLOW, 1 s
   "20_TANKS_IP_DATA_RIO_03_FIRST_TANK_BWT_LEVEL_HIHI" : Bool = PLC "20_TANKS_IP_DATA".RIO_03.FIRST_TANK.BWT_LEVEL_HIHI, 1 s
   "20_TANKS_IP_DATA_RIO_03_FIRST_TANK_GTT_ISOL_VALVE_OPEN" : Bool = PLC "20_TANKS_IP_DATA".RIO_03.FIRST_TANK.GTT_ISOL_VALVE_OPEN, 1 s
   "20_TANKS_IP_DATA_RIO_03_FIRST_TANK_GTT_ISOL_VALVE_CLSD" : Bool = PLC "20_TANKS_IP_DATA".RIO_03.FIRST_TANK.GTT_ISOL_VALVE_CLSD, 1 s
   "20_TANKS_IP_DATA_RIO_03_SECOND_TANK_BWT_LEVEL_HIHI" : Bool = PLC "20_TANKS_IP_DATA".RIO_03.SECOND_TANK.BWT_LEVEL_HIHI, 1 s
   "504_Tank Grouping_DB2020_RUN TANK 7" : Bool = PLC "504_Tank Grouping_DB2020"."RUN TANK 7", 1 s
   "20_TANKS_IP_DATA_RIO_03_SECOND_TANK_USD_FLOW" : Real = PLC "20_TANKS_IP_DATA".RIO_03.SECOND_TANK.USD_FLOW, 1 s
   "20_TANKS_IP_DATA_RIO_03_SECOND_TANK_MBG_FLOW" : Real = PLC "20_TANKS_IP_DATA".RIO_03.SECOND_TANK.MBG_FLOW, 1 s
   "20_TANKS_IP_DATA_RIO_03_SECOND_TANK_GTT_ISOL_VALVE_OPEN" : Bool = PLC "20_TANKS_IP_DATA".RIO_03.SECOND_TANK.GTT_ISOL_VALVE_OPEN, 1 s
   "20_TANKS_IP_DATA_RIO_03_SECOND_TANK_GTT_ISOL_VALVE_CLSD" : Bool = PLC "20_TANKS_IP_DATA".RIO_03.SECOND_TANK.GTT_ISOL_VALVE_CLSD, 1 s
   "20_TANKS_IP_DATA_RIO_04_FIRST_TANK_BWT_LEVEL_HIHI" : Bool = PLC "20_TANKS_IP_DATA".RIO_04.FIRST_TANK.BWT_LEVEL_HIHI, 1 s
   "20_TANKS_IP_DATA_RIO_04_FIRST_TANK_USD_FLOW" : Real = PLC "20_TANKS_IP_DATA".RIO_04.FIRST_TANK.USD_FLOW, 1 s
   "20_TANKS_IP_DATA_RIO_04_FIRST_TANK_MBG_FLOW" : Real = PLC "20_TANKS_IP_DATA".RIO_04.FIRST_TANK.MBG_FLOW, 1 s
   "20_TANKS_IP_DATA_RIO_04_FIRST_TANK_GTT_ISOL_VALVE_OPEN" : Bool = PLC "20_TANKS_IP_DATA".RIO_04.FIRST_TANK.GTT_ISOL_VALVE_OPEN, 1 s
   "20_TANKS_IP_DATA_RIO_04_FIRST_TANK_GTT_ISOL_VALVE_CLSD" : Bool = PLC "20_TANKS_IP_DATA".RIO_04.FIRST_TANK.GTT_ISOL_VALVE_CLSD, 1 s
   "20_TANKS_IP_DATA_RIO_04_SECOND_TANK_BWT_LEVEL_HIHI" : Bool = PLC "20_TANKS_IP_DATA".RIO_04.SECOND_TANK.BWT_LEVEL_HIHI, 1 s
   "20_TANKS_IP_DATA_RIO_04_SECOND_TANK_USD_FLOW" : Real = PLC "20_TANKS_IP_DATA".RIO_04.SECOND_TANK.USD_FLOW, 1 s
   "20_TANKS_IP_DATA_RIO_04_SECOND_TANK_MBG_FLOW" : Real = PLC "20_TANKS_IP_DATA".RIO_04.SECOND_TANK.MBG_FLOW, 1 s
   "20_TANKS_IP_DATA_RIO_04_SECOND_TANK_GTT_ISOL_VALVE_OPEN" : Bool = PLC "20_TANKS_IP_DATA".RIO_04.SECOND_TANK.GTT_ISOL_VALVE_OPEN, 1 s
   "20_TANKS_IP_DATA_RIO_04_SECOND_TANK_GTT_ISOL_VALVE_CLSD" : Bool = PLC "20_TANKS_IP_DATA".RIO_04.SECOND_TANK.GTT_ISOL_VALVE_CLSD, 1 s
   "20_TANKS_IP_DATA_RIO_05_FIRST_TANK_BWT_LEVEL_HIHI" : Bool = PLC "20_TANKS_IP_DATA".RIO_05.FIRST_TANK.BWT_LEVEL_HIHI, 1 s
   "20_TANKS_IP_DATA_RIO_05_FIRST_TANK_MBG_FLOW" : Real = PLC "20_TANKS_IP_DATA".RIO_05.FIRST_TANK.MBG_FLOW, 1 s
   "20_TANKS_IP_DATA_RIO_05_FIRST_TANK_USD_FLOW" : Real = PLC "20_TANKS_IP_DATA".RIO_05.FIRST_TANK.USD_FLOW, 1 s
   "20_TANKS_IP_DATA_RIO_05_FIRST_TANK_GTT_ISOL_VALVE_OPEN" : Bool = PLC "20_TANKS_IP_DATA".RIO_05.FIRST_TANK.GTT_ISOL_VALVE_OPEN, 1 s
   "20_TANKS_IP_DATA_RIO_05_FIRST_TANK_GTT_ISOL_VALVE_CLSD" : Bool = PLC "20_TANKS_IP_DATA".RIO_05.FIRST_TANK.GTT_ISOL_VALVE_CLSD, 1 s
   "20_TANKS_IP_DATA_RIO_05_SECOND_TANK_BWT_LEVEL_HIHI" : Bool = PLC "20_TANKS_IP_DATA".RIO_05.SECOND_TANK.BWT_LEVEL_HIHI, 1 s
   "20_TANKS_IP_DATA_RIO_05_SECOND_TANK_USD_FLOW" : Real = PLC "20_TANKS_IP_DATA".RIO_05.SECOND_TANK.USD_FLOW, 1 s
   "20_TANKS_IP_DATA_RIO_05_SECOND_TANK_MBG_FLOW" : Real = PLC "20_TANKS_IP_DATA".RIO_05.SECOND_TANK.MBG_FLOW, 1 s
   "20_TANKS_IP_DATA_RIO_05_SECOND_TANK_GTT_ISOL_VALVE_OPEN" : Bool = PLC "20_TANKS_IP_DATA".RIO_05.SECOND_TANK.GTT_ISOL_VALVE_OPEN, 1 s
   "20_TANKS_IP_DATA_RIO_05_SECOND_TANK_GTT_ISOL_VALVE_CLSD" : Bool = PLC "20_TANKS_IP_DATA".RIO_05.SECOND_TANK.GTT_ISOL_VALVE_CLSD, 1 s
   "20_TANKS_IP_DATA_RIO_06_FIRST_TANK_BWT_LEVEL_HIHI" : Bool = PLC "20_TANKS_IP_DATA".RIO_06.FIRST_TANK.BWT_LEVEL_HIHI, 1 s
   "20_TANKS_IP_DATA_RIO_06_FIRST_TANK_USD_FLOW" : Real = PLC "20_TANKS_IP_DATA".RIO_06.FIRST_TANK.USD_FLOW, 1 s
   "20_TANKS_IP_DATA_RIO_06_FIRST_TANK_MBG_FLOW" : Real = PLC "20_TANKS_IP_DATA".RIO_06.FIRST_TANK.MBG_FLOW, 1 s
   "20_TANKS_IP_DATA_RIO_06_FIRST_TANK_GTT_ISOL_VALVE_OPEN" : Bool = PLC "20_TANKS_IP_DATA".RIO_06.FIRST_TANK.GTT_ISOL_VALVE_OPEN, 1 s
   "20_TANKS_IP_DATA_RIO_06_FIRST_TANK_GTT_ISOL_VALVE_CLSD" : Bool = PLC "20_TANKS_IP_DATA".RIO_06.FIRST_TANK.GTT_ISOL_VALVE_CLSD, 1 s
   "20_TANKS_IP_DATA_RIO_06_SECOND_TANK_BWT_LEVEL_HIHI" : Bool = PLC "20_TANKS_IP_DATA".RIO_06.SECOND_TANK.BWT_LEVEL_HIHI, 1 s
   "20_TANKS_IP_DATA_RIO_06_SECOND_TANK_USD_FLOW" : Real = PLC "20_TANKS_IP_DATA".RIO_06.SECOND_TANK.USD_FLOW, 1 s
   "20_TANKS_IP_DATA_RIO_06_SECOND_TANK_MBG_FLOW" : Real = PLC "20_TANKS_IP_DATA".RIO_06.SECOND_TANK.MBG_FLOW, 1 s
   "20_TANKS_IP_DATA_RIO_06_SECOND_TANK_GTT_ISOL_VALVE_OPEN" : Bool = PLC "20_TANKS_IP_DATA".RIO_06.SECOND_TANK.GTT_ISOL_VALVE_OPEN, 1 s
   "20_TANKS_IP_DATA_RIO_06_SECOND_TANK_GTT_ISOL_VALVE_CLSD" : Bool = PLC "Sequence Times_DB"."Re-Ox Timer"."Minutes Left", 1 s
   "20_TANKS_IP_DATA_RIO_07_FIRST_TANK_BWT_LEVEL_HIHI" : Bool = PLC "20_TANKS_IP_DATA".RIO_07.FIRST_TANK.BWT_LEVEL_HIHI, 1 s
   "20_TANKS_IP_DATA_RIO_07_FIRST_TANK_GTT_ISOL_VALVE_OPEN" : Bool = PLC "20_TANKS_IP_DATA".RIO_07.FIRST_TANK.GTT_ISOL_VALVE_OPEN, 1 s
   "20_TANKS_IP_DATA_RIO_07_FIRST_TANK_GTT_ISOL_VALVE_CLSD" : Bool = PLC "20_TANKS_IP_DATA".RIO_07.FIRST_TANK.GTT_ISOL_VALVE_CLSD, 1 s